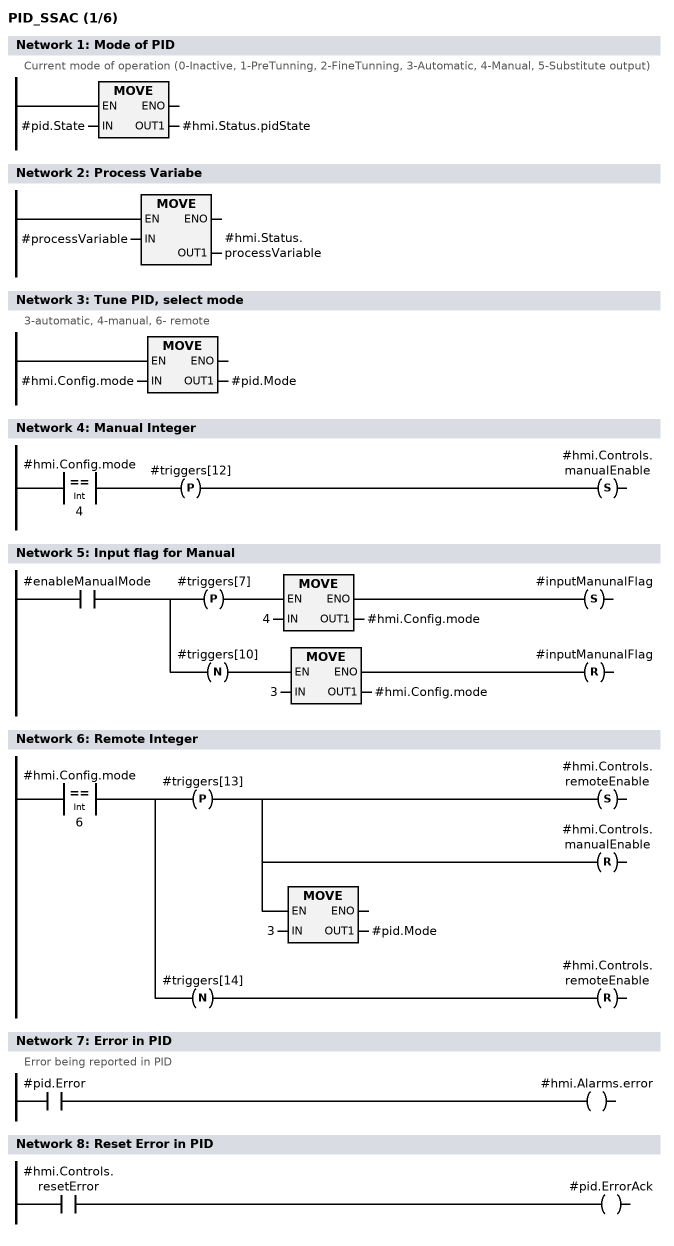
   RUNG wire#powerrail
      Move(in := #pid.State, out1 => #hmi.Status.pidState)
   END_RUNG
   // the same network as SCL:
   #hmi.Status.pidState := #pid.State;
END_REGION

REGION Network 2: Process Variabe
   RUNG wire#powerrail
      Move(in := #processVariable, out1 => #hmi.Status.processVariable)
   END_RUNG
   // the same network as SCL:
   #hmi.Status.processVariable := #processVariable;
END_REGION

REGION Network 3: Tune PID, select mode
   // 3-automatic, 4-manual, 6- remote
   RUNG wire#powerrail
      Move(in := #hmi.Config.mode, out1 => #pid.Mode)
   END_RUNG
   // the same network as SCL:
   #pid.Mode := #hmi.Config.mode;
END_REGION

REGION Network 4: Manual Integer
   RUNG wire#powerrail
      { S7_Templates := "SrcType := Int" } EQ_Contact(in1 := #hmi.Config.mode, in2 := 4)
      P_Trig( #triggers[12] )
      S_Coil( #hmi.Controls.manualEnable )
   END_RUNG
   // the same network as SCL:
   #_w1 := #hmi.Config.mode = 4;
   #_w2 := #_w1 AND NOT #triggers[12];   // rising edge
   #triggers[12] := #_w1;
   IF #_w2 THEN #hmi.Controls.manualEnable := TRUE; END_IF;
END_REGION

REGION Network 5: Input flag for Manual
   RUNG wire#powerrail
      Contact( #enableManualMode )
      wire#w1
      P_Trig( #triggers[7] )
      Move(in := 4, out1 => #hmi.Config.mode)
      S_Coil( #inputManunalFlag )
   END_RUNG
   RUNG wire#w1
      N_Trig( #triggers[10] )
      Move(in := 3, out1 => #hmi.Config.mode)
      R_Coil( #inputManunalFlag )
   END_RUNG
   // the same network as SCL:
   #_w1 := #enableManualMode AND NOT #triggers[7];   // rising edge
   #triggers[7] := #enableManualMode;
   IF #_w1 THEN
       #hmi.Config.mode := 4;
       #inputManunalFlag := TRUE;
   END_IF;
   #_w2 := NOT #enableManualMode AND #triggers[10];   // falling edge
   #triggers[10] := #enableManualMode;
   IF #_w2 THEN
       #hmi.Config.mode := 3;
       #inputManunalFlag := FALSE;
   END_IF;
END_REGION

REGION Network 6: Remote Integer
   RUNG wire#powerrail
      { S7_Templates := "SrcType := Int" } EQ_Contact(in1 := #hmi.Config.mode, in2 := 6)
      wire#w1
      P_Trig( #triggers[13] )
      wire#w2
      S_Coil( #hmi.Controls.remoteEnable )
   END_RUNG
   RUNG wire#w2
      R_Coil( #hmi.Controls.manualEnable )
   END_RUNG
   RUNG wire#w2
      Move(in := 3, out1 => #pid.Mode)
   END_RUNG
   RUNG wire#w1
      N_Trig( #triggers[14] )
      R_Coil( #hmi.Controls.remoteEnable )
   END_RUNG
   // the same network as SCL:
   #_w1 := #hmi.Config.mode = 6;
   #_w2 := #_w1 AND NOT #triggers[13];   // rising edge
   #triggers[13] := #_w1;
   IF #_w2 THEN
       #hmi.Controls.remoteEnable := TRUE;
       #hmi.Controls.manualEnable := FALSE;
       #pid.Mode := 3;
   END_IF;
   #_w3 := NOT #_w1 AND #triggers[14];   // falling edge
   #triggers[14] := #_w1;
   IF #_w3 THEN #hmi.Controls.remoteEnable := FALSE; END_IF;
END_REGION

REGION Network 7: Error in PID
   // Error being reported in PID
   RUNG wire#powerrail
      Contact( #pid.Error )
      Coil( #hmi.Alarms.error )
   END_RUNG
   // the same network as SCL:
   #hmi.Alarms.error := #pid.Error;
END_REGION

REGION Network 8: Reset Error in PID
   RUNG wire#powerrail
      Contact( #hmi.Controls.resetError )
      Coil( #pid.ErrorAck )
   END_RUNG
   // the same network as SCL:
   #pid.ErrorAck := #hmi.Controls.resetError;
END_REGION

REGION Network 9: Reset the controller if a change of Mode has been requested
   // mode 2 3 4 available thru here
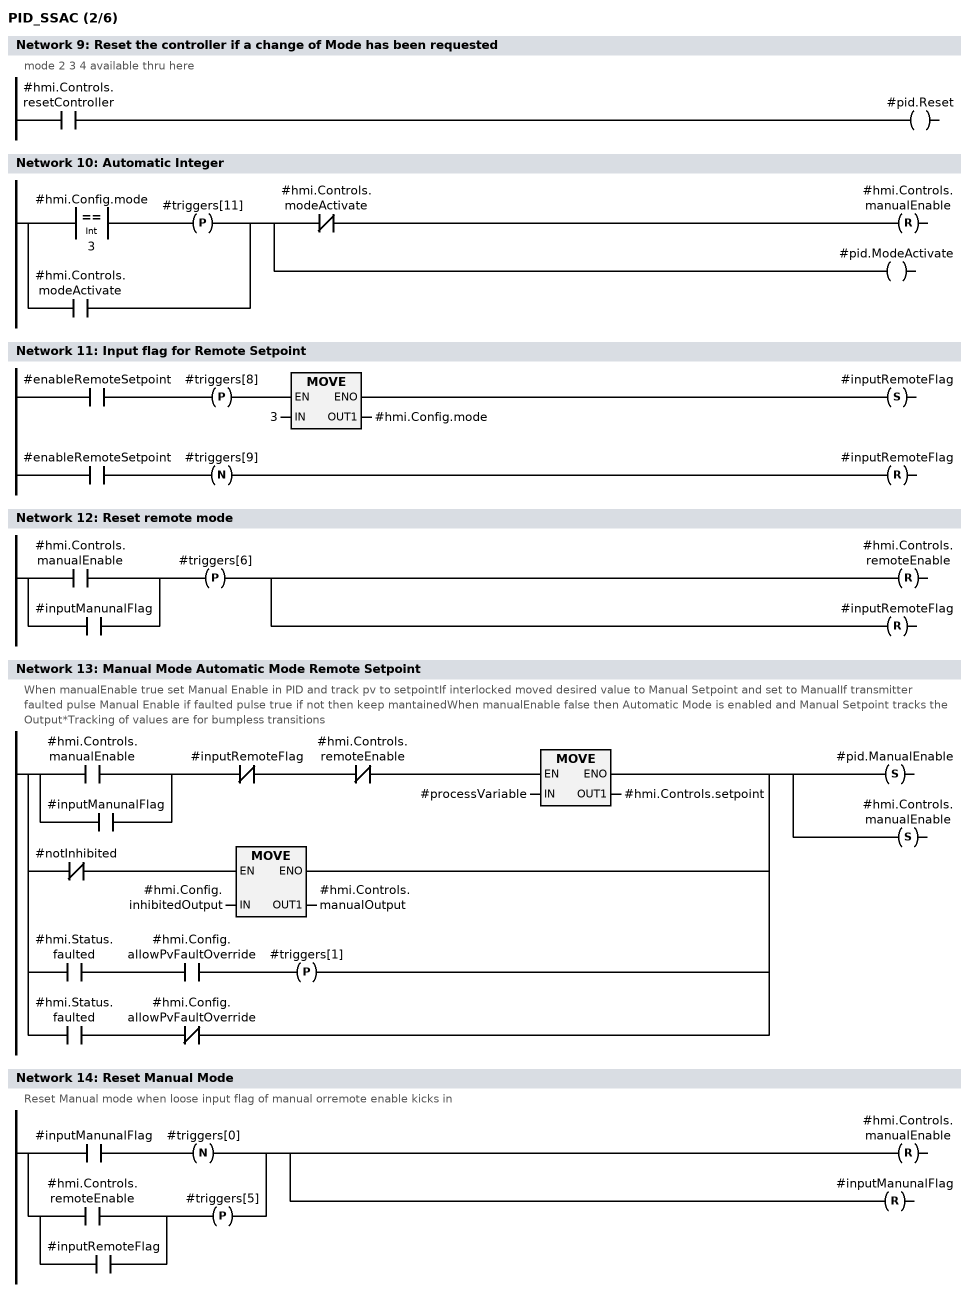
   RUNG wire#powerrail
      Contact( #hmi.Controls.resetController )
      Coil( #pid.Reset )
   END_RUNG
   // the same network as SCL:
   #pid.Reset := #hmi.Controls.resetController;
END_REGION

REGION Network 10: Automatic Integer
   RUNG wire#powerrail
      { S7_Templates := "SrcType := Int" } EQ_Contact(in1 := #hmi.Config.mode, in2 := 3)
      P_Trig( #triggers[11] )
      wire#w1
      I_Contact( #hmi.Controls.modeActivate )
      R_Coil( #hmi.Controls.manualEnable )
   END_RUNG
   RUNG wire#powerrail
      Contact( #hmi.Controls.modeActivate )
   END_RUNG wire#w1
   RUNG wire#w1
      Coil( #pid.ModeActivate )
   END_RUNG
   // the same network as SCL:
   #_w1 := #hmi.Config.mode = 3;
   #_w2 := #_w1 AND NOT #triggers[11];   // rising edge
   #triggers[11] := #_w1;
   #_w3 := #_w2 OR #hmi.Controls.modeActivate;
   IF #_w3 AND NOT #hmi.Controls.modeActivate THEN #hmi.Controls.manualEnable := FALSE; END_IF;
   #pid.ModeActivate := #_w3;
END_REGION

REGION Network 11: Input flag for Remote Setpoint
   RUNG wire#powerrail
      Contact( #enableRemoteSetpoint )
      P_Trig( #triggers[8] )
      Move(in := 3, out1 => #hmi.Config.mode)
      S_Coil( #inputRemoteFlag )
   END_RUNG
   RUNG wire#powerrail
      Contact( #enableRemoteSetpoint )
      N_Trig( #triggers[9] )
      R_Coil( #inputRemoteFlag )
   END_RUNG
   // the same network as SCL:
   #_w1 := #enableRemoteSetpoint AND NOT #triggers[8];   // rising edge
   #triggers[8] := #enableRemoteSetpoint;
   IF #_w1 THEN
       #hmi.Config.mode := 3;
       #inputRemoteFlag := TRUE;
   END_IF;
   #_w2 := NOT #enableRemoteSetpoint AND #triggers[9];   // falling edge
   #triggers[9] := #enableRemoteSetpoint;
   IF #_w2 THEN #inputRemoteFlag := FALSE; END_IF;
END_REGION

REGION Network 12: Reset remote mode
   RUNG wire#powerrail
      Contact( #hmi.Controls.manualEnable )
      wire#w1
      P_Trig( #triggers[6] )
      wire#w2
      R_Coil( #hmi.Controls.remoteEnable )
   END_RUNG
   RUNG wire#powerrail
      Contact( #inputManunalFlag )
   END_RUNG wire#w1
   RUNG wire#w2
      R_Coil( #inputRemoteFlag )
   END_RUNG
   // the same network as SCL:
   #_w1 := #hmi.Controls.manualEnable OR #inputManunalFlag;
   #_w2 := #_w1 AND NOT #triggers[6];   // rising edge
   #triggers[6] := #_w1;
   IF #_w2 THEN
       #hmi.Controls.remoteEnable := FALSE;
       #inputRemoteFlag := FALSE;
   END_IF;
END_REGION

REGION Network 13: Manual Mode Automatic Mode Remote Setpoint
   // When manualEnable true set Manual Enable in PID and track pv to setpointIf interlocked moved desired value to Manual Setpoint and set to ManualIf transmitter faulted pulse Manual Enable if faulted pulse true if not then keep mantainedWhen manualEnable false then Automatic Mode is enabled and Manual Setpoint tracks the Output*Tracking of values are for bumpless transitions
   RUNG wire#powerrail
      Contact( #hmi.Controls.manualEnable )
      wire#w1
      I_Contact( #inputRemoteFlag )
      I_Contact( #hmi.Controls.remoteEnable )
      Move(in := #processVariable, out1 => #hmi.Controls.setpoint)
      wire#w2
      S_Coil( #pid.ManualEnable )
   END_RUNG
   RUNG wire#powerrail
      Contact( #inputManunalFlag )
   END_RUNG wire#w1
   RUNG wire#powerrail
      I_Contact( #notInhibited )
      Move(in := #hmi.Config.inhibitedOutput, out1 => #hmi.Controls.manualOutput)
   END_RUNG wire#w2
   RUNG wire#powerrail
      Contact( #hmi.Status.faulted )
      Contact( #hmi.Config.allowPvFaultOverride )
      P_Trig( #triggers[1] )
   END_RUNG wire#w2
   RUNG wire#powerrail
      Contact( #hmi.Status.faulted )
      I_Contact( #hmi.Config.allowPvFaultOverride )
   END_RUNG wire#w2
   RUNG wire#w2
      S_Coil( #hmi.Controls.manualEnable )
   END_RUNG
   // the same network as SCL:
   #_w1 := (#hmi.Controls.manualEnable OR #inputManunalFlag) AND NOT #inputRemoteFlag AND NOT #hmi.Controls.remoteEnable;
   IF #_w1 THEN #hmi.Controls.setpoint := #processVariable; END_IF;
   IF NOT #notInhibited THEN #hmi.Controls.manualOutput := #hmi.Config.inhibitedOutput; END_IF;
   #_w2 := #hmi.Status.faulted AND #hmi.Config.allowPvFaultOverride;
   #_w3 := #_w2 AND NOT #triggers[1];   // rising edge
   #triggers[1] := #_w2;
   IF #_w1 OR NOT #notInhibited OR #_w3 OR (#hmi.Status.faulted AND NOT #hmi.Config.allowPvFaultOverride) THEN
       #pid.ManualEnable := TRUE;
       #hmi.Controls.manualEnable := TRUE;
   END_IF;
END_REGION

REGION Network 14: Reset Manual Mode
   // Reset Manual mode when loose input flag of manual orremote enable kicks in
   RUNG wire#powerrail
      Contact( #inputManunalFlag )
      N_Trig( #triggers[0] )
      wire#w1
      R_Coil( #hmi.Controls.manualEnable )
   END_RUNG
   RUNG wire#powerrail
      Contact( #hmi.Controls.remoteEnable )
      wire#w2
      P_Trig( #triggers[5] )
   END_RUNG wire#w1
   RUNG wire#powerrail
      Contact( #inputRemoteFlag )
   END_RUNG wire#w2
   RUNG wire#w1
      R_Coil( #inputManunalFlag )
   END_RUNG
   // the same network as SCL:
   #_w1 := NOT #inputManunalFlag AND #triggers[0];   // falling edge
   #triggers[0] := #inputManunalFlag;
   #_w2 := #hmi.Controls.remoteEnable OR #inputRemoteFlag;
   #_w3 := #_w2 AND NOT #triggers[5];   // rising edge
   #triggers[5] := #_w2;
   IF #_w1 OR #_w3 THEN
       #hmi.Controls.manualEnable := FALSE;
       #inputManunalFlag := FALSE;
   END_IF;
END_REGION

REGION Network 15: Automatic Mode
   // IF not in manual and not in remote then in Automatic mode, reset Manual Mode of  PID
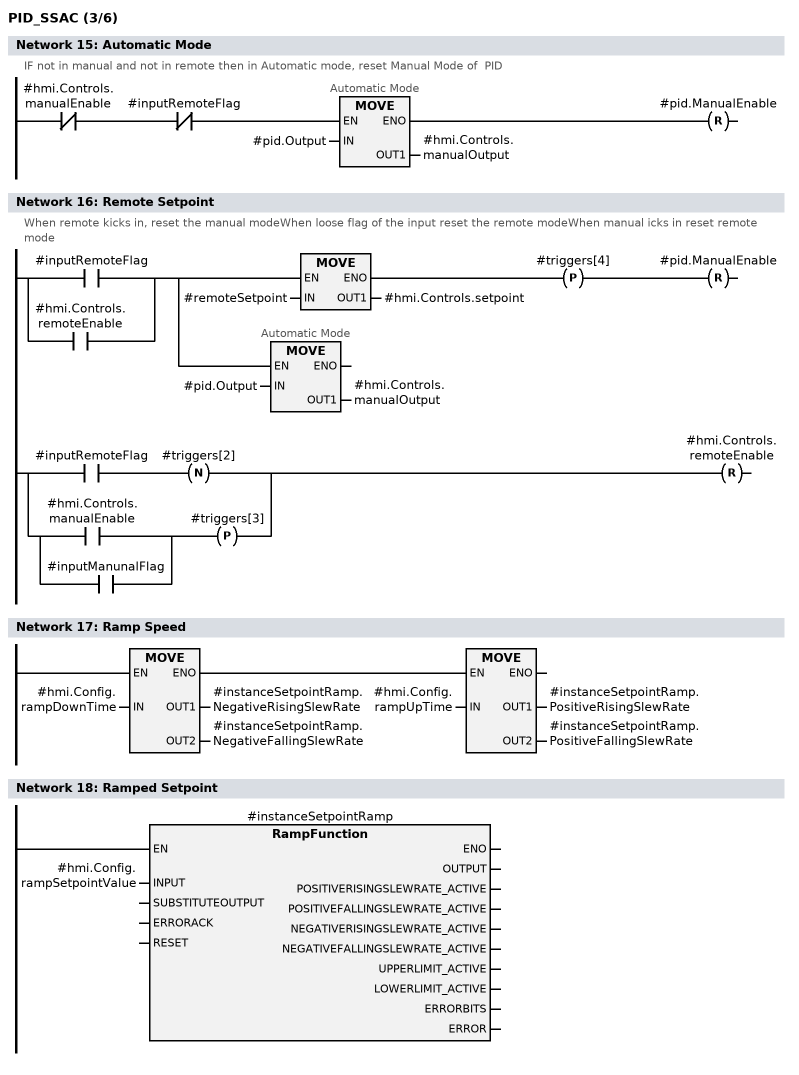
   RUNG wire#powerrail
      I_Contact( #hmi.Controls.manualEnable )
      I_Contact( #inputRemoteFlag )
      Move(in := #pid.Output, out1 => #hmi.Controls.manualOutput)   // Automatic Mode
      R_Coil( #pid.ManualEnable )
   END_RUNG
   // the same network as SCL:
   IF NOT #hmi.Controls.manualEnable AND NOT #inputRemoteFlag THEN
       #hmi.Controls.manualOutput := #pid.Output;   // Automatic Mode
       #pid.ManualEnable := FALSE;
   END_IF;
END_REGION

REGION Network 16: Remote Setpoint
   // When remote kicks in, reset the manual modeWhen loose flag of the input reset the remote modeWhen manual icks in reset remote mode
   RUNG wire#powerrail
      Contact( #inputRemoteFlag )
      wire#w1
      Move(in := #remoteSetpoint, out1 => #hmi.Controls.setpoint)
      P_Trig( #triggers[4] )
      R_Coil( #pid.ManualEnable )
   END_RUNG
   RUNG wire#powerrail
      Contact( #hmi.Controls.remoteEnable )
   END_RUNG wire#w1
   RUNG wire#w1
      Move(in := #pid.Output, out1 => #hmi.Controls.manualOutput)   // Automatic Mode
   END_RUNG
   RUNG wire#powerrail
      Contact( #inputRemoteFlag )
      N_Trig( #triggers[2] )
      wire#w2
      R_Coil( #hmi.Controls.remoteEnable )
   END_RUNG
   RUNG wire#powerrail
      Contact( #hmi.Controls.manualEnable )
      wire#w3
      P_Trig( #triggers[3] )
   END_RUNG wire#w2
   RUNG wire#powerrail
      Contact( #inputManunalFlag )
   END_RUNG wire#w3
   // the same network as SCL:
   #_w1 := #inputRemoteFlag OR #hmi.Controls.remoteEnable;
   IF #_w1 THEN #hmi.Controls.setpoint := #remoteSetpoint; END_IF;
   #_w2 := #_w1 AND NOT #triggers[4];   // rising edge
   #triggers[4] := #_w1;
   IF #_w2 THEN #pid.ManualEnable := FALSE; END_IF;
   IF #_w1 THEN
       #hmi.Controls.manualOutput := #pid.Output;   // Automatic Mode
   END_IF;
   #_w3 := NOT #inputRemoteFlag AND #triggers[2];   // falling edge
   #triggers[2] := #inputRemoteFlag;
   #_w4 := #hmi.Controls.manualEnable OR #inputManunalFlag;
   #_w5 := #_w4 AND NOT #triggers[3];   // rising edge
   #triggers[3] := #_w4;
   IF #_w3 OR #_w5 THEN #hmi.Controls.remoteEnable := FALSE; END_IF;
END_REGION

REGION Network 17: Ramp Speed
   RUNG wire#powerrail
      Move(in := #hmi.Config.rampDownTime, out1 => #instanceSetpointRamp.NegativeRisingSlewRate, out2 => #instanceSetpointRamp.NegativeFallingSlewRate)
      Move(in := #hmi.Config.rampUpTime, out1 => #instanceSetpointRamp.PositiveRisingSlewRate, out2 => #instanceSetpointRamp.PositiveFallingSlewRate)
   END_RUNG
   // the same network as SCL:
   #instanceSetpointRamp.NegativeRisingSlewRate := #hmi.Config.rampDownTime;
   #instanceSetpointRamp.NegativeFallingSlewRate := #hmi.Config.rampDownTime;
   #instanceSetpointRamp.PositiveRisingSlewRate := #hmi.Config.rampUpTime;
   #instanceSetpointRamp.PositiveFallingSlewRate := #hmi.Config.rampUpTime;
END_REGION

REGION Network 18: Ramped Setpoint
   #instanceSetpointRamp(Input := #hmi.Config.rampSetpointValue);   // RampFunction
END_REGION

REGION Network 19: Setpoint Control
   // If ramp enabled then move ramped setpointif ramp disabled then move hmi setpoint
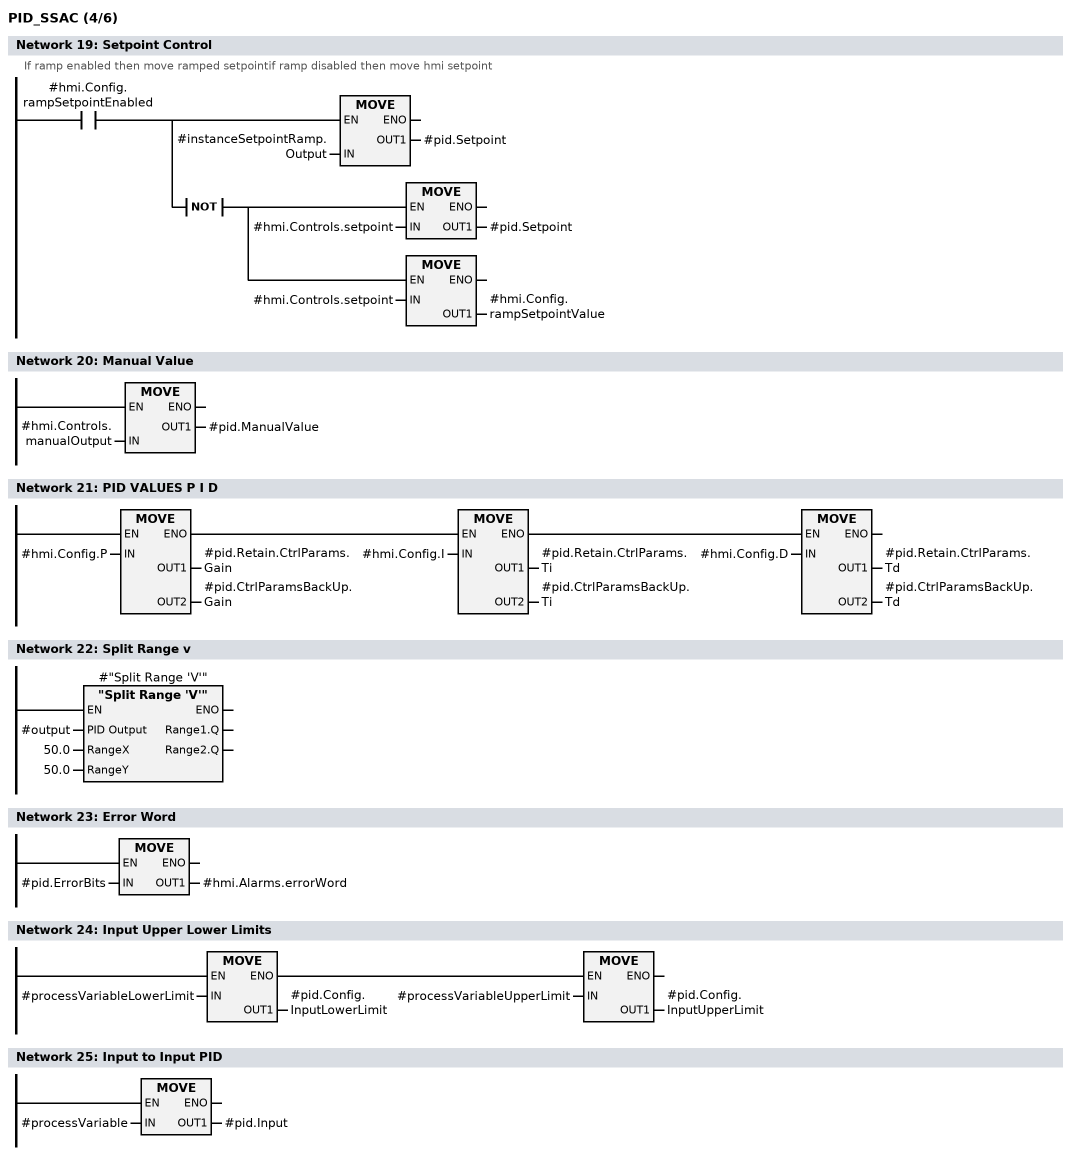
   RUNG wire#powerrail
      Contact( #hmi.Config.rampSetpointEnabled )
      wire#w1
      Move(in := #instanceSetpointRamp.Output, out1 => #pid.Setpoint)
   END_RUNG
   RUNG wire#w1
      Not()
      wire#w2
      Move(in := #hmi.Controls.setpoint, out1 => #pid.Setpoint)
   END_RUNG
   RUNG wire#w2
      Move(in := #hmi.Controls.setpoint, out1 => #hmi.Config.rampSetpointValue)
   END_RUNG
   // the same network as SCL:
   IF #hmi.Config.rampSetpointEnabled THEN #pid.Setpoint := #instanceSetpointRamp.Output; END_IF;
   IF NOT #hmi.Config.rampSetpointEnabled THEN
       #pid.Setpoint := #hmi.Controls.setpoint;
       #hmi.Config.rampSetpointValue := #hmi.Controls.setpoint;
   END_IF;
END_REGION

REGION Network 20: Manual Value
   RUNG wire#powerrail
      Move(in := #hmi.Controls.manualOutput, out1 => #pid.ManualValue)
   END_RUNG
   // the same network as SCL:
   #pid.ManualValue := #hmi.Controls.manualOutput;
END_REGION

REGION Network 21: PID VALUES P I D
   RUNG wire#powerrail
      Move(in := #hmi.Config.P, out1 => #pid.Retain.CtrlParams.Gain, out2 => #pid.CtrlParamsBackUp.Gain)
      Move(in := #hmi.Config.I, out1 => #pid.Retain.CtrlParams.Ti, out2 => #pid.CtrlParamsBackUp.Ti)
      Move(in := #hmi.Config.D, out1 => #pid.Retain.CtrlParams.Td, out2 => #pid.CtrlParamsBackUp.Td)
   END_RUNG
   // the same network as SCL:
   #pid.Retain.CtrlParams.Gain := #hmi.Config.P;
   #pid.CtrlParamsBackUp.Gain := #hmi.Config.P;
   #pid.Retain.CtrlParams.Ti := #hmi.Config.I;
   #pid.CtrlParamsBackUp.Ti := #hmi.Config.I;
   #pid.Retain.CtrlParams.Td := #hmi.Config.D;
   #pid.CtrlParamsBackUp.Td := #hmi.Config.D;
END_REGION

REGION Network 22: Split Range v
   RUNG wire#powerrail
      #"Split Range 'V'"("PID Output" := #output, RangeX := 50.0, RangeY := 50.0, "Range1.Q" =>, "Range2.Q" =>)
   END_RUNG
   // the same network as SCL:
   #"Split Range 'V'"("PID Output" := #output, RangeX := 50.0, RangeY := 50.0);   // "Split Range 'V'"
END_REGION

REGION Network 23: Error Word
   RUNG wire#powerrail
      Move(in := #pid.ErrorBits, out1 => #hmi.Alarms.errorWord)
   END_RUNG
   // the same network as SCL:
   #hmi.Alarms.errorWord := #pid.ErrorBits;
END_REGION

REGION Network 24: Input Upper Lower Limits
   RUNG wire#powerrail
      Move(in := #processVariableLowerLimit, out1 => #pid.Config.InputLowerLimit)
      Move(in := #processVariableUpperLimit, out1 => #pid.Config.InputUpperLimit)
   END_RUNG
   // the same network as SCL:
   #pid.Config.InputLowerLimit := #processVariableLowerLimit;
   #pid.Config.InputUpperLimit := #processVariableUpperLimit;
END_REGION

REGION Network 25: Input to Input PID
   RUNG wire#powerrail
      Move(in := #processVariable, out1 => #pid.Input)
   END_RUNG
   // the same network as SCL:
   #pid.Input := #processVariable;
END_REGION

REGION Network 26: Outputs
   // Outputs of PID block
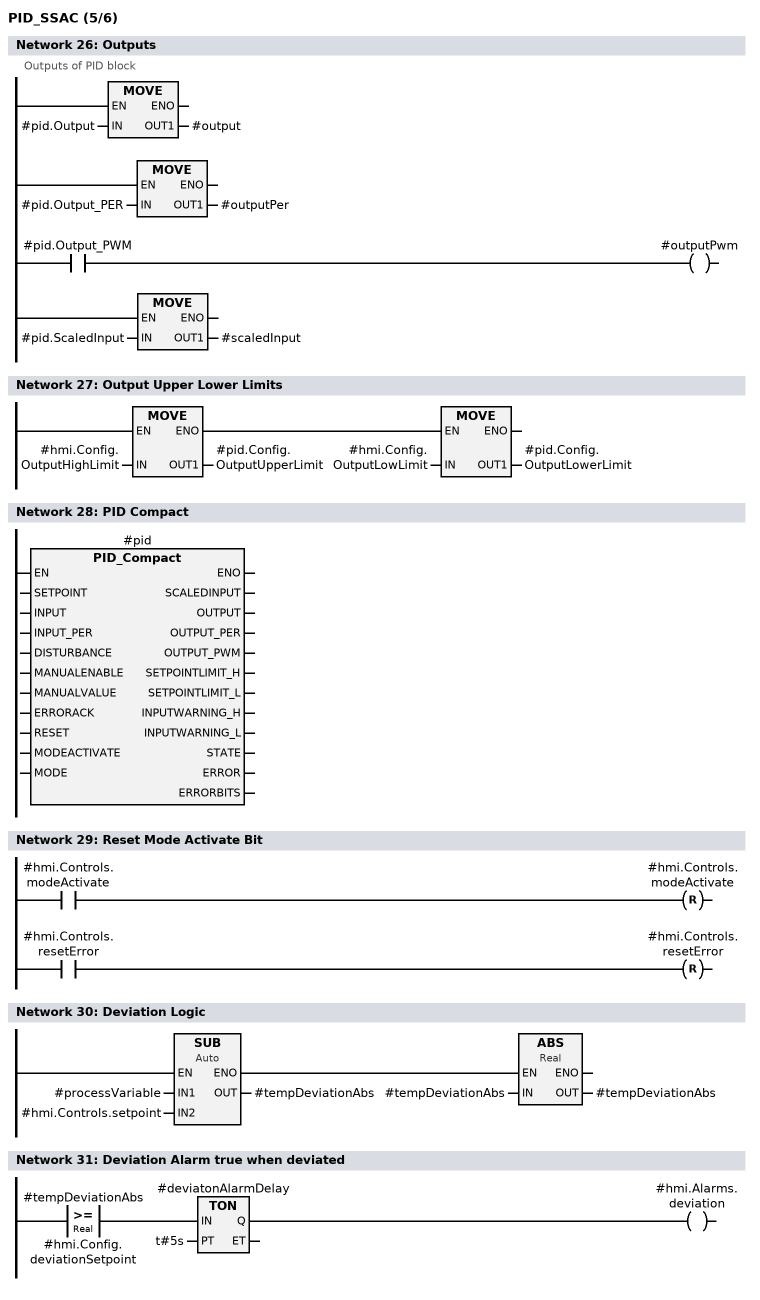
   RUNG wire#powerrail
      Move(in := #pid.Output, out1 => #output)
   END_RUNG
   RUNG wire#powerrail
      Move(in := #pid.Output_PER, out1 => #outputPer)
   END_RUNG
   RUNG wire#powerrail
      Contact( #pid.Output_PWM )
      Coil( #outputPwm )
   END_RUNG
   RUNG wire#powerrail
      Move(in := #pid.ScaledInput, out1 => #scaledInput)
   END_RUNG
   // the same network as SCL:
   #output := #pid.Output;
   #outputPer := #pid.Output_PER;
   #outputPwm := #pid.Output_PWM;
   #scaledInput := #pid.ScaledInput;
END_REGION

REGION Network 27: Output Upper Lower Limits
   RUNG wire#powerrail
      Move(in := #hmi.Config.OutputHighLimit, out1 => #pid.Config.OutputUpperLimit)
      Move(in := #hmi.Config.OutputLowLimit, out1 => #pid.Config.OutputLowerLimit)
   END_RUNG
   // the same network as SCL:
   #pid.Config.OutputUpperLimit := #hmi.Config.OutputHighLimit;
   #pid.Config.OutputLowerLimit := #hmi.Config.OutputLowLimit;
END_REGION

REGION Network 28: PID Compact
   #pid();   // PID_Compact
END_REGION

REGION Network 29: Reset Mode Activate Bit
   RUNG wire#powerrail
      Contact( #hmi.Controls.modeActivate )
      R_Coil( #hmi.Controls.modeActivate )
   END_RUNG
   RUNG wire#powerrail
      Contact( #hmi.Controls.resetError )
      R_Coil( #hmi.Controls.resetError )
   END_RUNG
   // the same network as SCL:
   IF #hmi.Controls.modeActivate THEN #hmi.Controls.modeActivate := FALSE; END_IF;
   IF #hmi.Controls.resetError THEN #hmi.Controls.resetError := FALSE; END_IF;
END_REGION

REGION Network 30: Deviation Logic
   RUNG wire#powerrail
      Sub(in1 := #processVariable, in2 := #hmi.Controls.setpoint, out => #tempDeviationAbs)
      { S7_Templates := "SrcType := Real" } Abs(in := #tempDeviationAbs, out => #tempDeviationAbs)
   END_RUNG
   // the same network as SCL:
   #tempDeviationAbs := #processVariable - #hmi.Controls.setpoint;
   #tempDeviationAbs := ABS(#tempDeviationAbs);
END_REGION

REGION Network 31: Deviation Alarm true when deviated
   #deviatonAlarmDelay(IN := #tempDeviationAbs >= #hmi.Config.deviationSetpoint, PT := t#5s);   // TON
   #hmi.Alarms.deviation := #deviatonAlarmDelay.Q;
END_REGION

REGION Network 32: PID inhibited (interlocked, off)
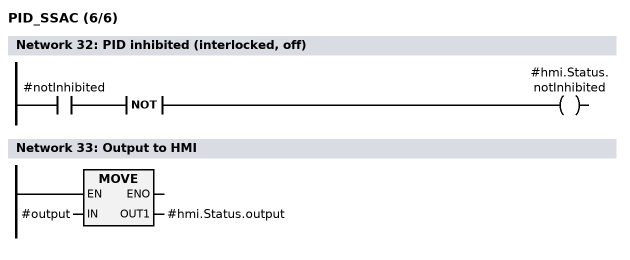
   RUNG wire#powerrail
      Contact( #notInhibited )
      Not()
      Coil( #hmi.Status.notInhibited )
   END_RUNG
   // the same network as SCL:
   #hmi.Status.notInhibited := NOT #notInhibited;
END_REGION

REGION Network 33: Output to HMI
   RUNG wire#powerrail
      Move(in := #output, out1 => #hmi.Status.output)
   END_RUNG
   // the same network as SCL:
   #hmi.Status.output := #output;
END_REGION
END_FUNCTION_BLOCK

FUNCTION_BLOCK "Totalizer_Siemens"   // FB3, SCL
{ S7_Optimized_Access := 'TRUE' }
VERSION : 0.1
   VAR_INPUT
      value : Real;
      intervall : Time;
      cycle : Time;
      reset : Bool;
   END_VAR
   VAR_OUTPUT
      total : Real;
   END_VAR
   VAR
      statAccum : Real;
   END_VAR
   VAR_TEMP
      tempIntervall : Real;
      tempCycle : Real;
      tempIntervallDInt : DInt;
      tempCycleDInt : DInt;
   END_VAR
BEGIN
   //Ist der Signalzustand der Variable "Reset" gleich True, so werden die Variablen
   //"Accum" und "Total" auf Null zurückgesetzt und es erfolgt keine Berechnung.
   //Beim Signalzustand False erfolgt zunächst eine Datentypumwandlung nach Real der beiden
   //Eingangsvariablen "Intervall" und "Cycle". Zuerst mit der Konvertierung von Time nach
   //DInt und anschließend von DInt nach Real.
   //Innerhalb eines Zyklus wird der Eingangswert der Variablen "Value" mit dem Wert der temporären Variablen
   //"Cycle_real" multipliziert und mit dem Wert der temporären Variablen "Intervall_real" dividiert.
   //Das Ergebnis wird anschließend in den Zwischenspeicher "Accum" abgelegt. Somit wird innerhalb eines jeden
   //Zykluses das Zwischenergebnis im "Accum" um diesen Wert inkrementiert, welches auch in jedem Zyklus zur
   //Ausgangsvariable "Total" transferiert wird.
   //***************************************************************************
   //If the signal status of the variable "Reset" is true, the variables "Accum" and "Total"
   //are set to zero and there is no calculation.
   //If the signal status is false, there is first a data type change to real of the two
   //input variables "Intervall" and "Cycle. After conversion from Time to DInit and from DInt to Real.
   //In a #Cycle the input #Value of the variable "Value" is multiplied by the #Value of the temporary variable
   //"Cycle_real" and then divided by the #Value of the temporary variable "Intervall_real". The result is then
   //stored in the buffer "Accum". This in one particular #Cycle the result in the "Accum" buffer is
   //incremented this #Value, which is also transferred to the output variable "Total" in that #Cycle too.

   IF #reset = true THEN
       #statAccum := 0.000000e000; //Die Variablen werden zurückgesetzt.
       #total := 0.000000e000; //The variables will be set to zero.
   ELSE
       #tempIntervallDInt := TIME_TO_DINT(#intervall);
       #tempIntervall := DINT_TO_REAL(#tempIntervallDInt);
       #tempCycleDInt := TIME_TO_DINT(#cycle);
       #tempCycle := DINT_TO_REAL(#tempCycleDInt);
       #statAccum := ((#value * #tempCycle) / #tempIntervall) + #statAccum;
       #total := #statAccum; //Kopiere Ergebnis nach #Total / Copy result to #Total.
   END_IF;
END_FUNCTION_BLOCK

FUNCTION_BLOCK "PID_TIA"   // FB814, LAD
{ S7_Optimized_Access := 'TRUE' }
VERSION : 0.1
   VAR_INPUT
      processVariable : Real;
      processVariableLowerLimit : Real;
      processVariableUpperLimit : Real;
      notInhibited : Bool := TRUE;
      remoteSetpoint : Real;
      enableManualMode : Bool;
      enableRemoteSetpoint : Bool;
   END_VAR
   VAR_OUTPUT
      scaledInput : Real;
      output : Real;   // Manipulated Value REAL
      outputPer : Int;   // Manipulated Value INT
      outputPwm : Bool;   // Output PWM
   END_VAR
   VAR_IN_OUT
      pid : PID_Compact;
   END_VAR
   VAR
      hmi : Struct
         Controls : Struct
            setpoint : Real;   // Setpoint sent to PID
            manualEnable : Bool;   // Enables Manual mode
            manualOutput : Real;   // Manual Output sent to PID 0 to 100 %
            remoteEnable : Bool;
            resetController : Bool;   // Resets Controller sent to PID
            resetError : Bool;   // ErrorAck to PID
            modeActivate : Bool;   // Execute the change of mode
         END_STRUCT;
         Config : Struct
            P : Real := 0.1;   // Proportional Control sent to PID
            I : Real := 10.0;   // Integral Control sent to PID
            D : Real := 0.0;   // Derivative Control sent to PID
            OutputHighLimit : Real := 100.0;   // Output Upper Limit sent to PID
            OutputLowLimit : Real := 0.0;   // Output Lower Limit sent to PID
            rampDownTime : Real := 1.0;
            rampUpTime : Real := 1.0;
            allowPvFaultOverride : Bool;   // Allows operator to override PV fault
            rampSetpointEnabled : Bool;   // Enables the ramping of a setpoint inside the PID
            rampSetpointValue : Real;   // Value to be reached in the ramp
            inhibitedOutput : Real := 0.0;   // Inhibited Value set by the Operator 0 to 100
            mode : Int := 4;   // Mode selected by operator 1=pretune,2=finetuning,3=automatic,4-manual, 5-Substitute output, 6-Remote
            enablePVtracking : Bool;
         END_STRUCT;
         Status : Struct
            faulted : Bool;   // Transmitter Faulted
            notInhibited : Bool;   // PID inhibited (interlocked, off)
            pidState : Int;   // Current mode of operation (0-Inactive, 1-SUT, 2-TIR, 3-Automatic, 4-Manual, 5-Substitute output)
            Output : Real;   // Output of the PID
         END_STRUCT;
         Alarms : Struct
            errorWord : DWord;   // Error Word of PID
            error : Bool;   // Error in PID
         END_STRUCT;
      END_STRUCT;
      triggers : Array[0..20] of Bool;
      inputManunalFlag : Bool;
      inputRemoteFlag : Bool;
      "Dont Overwrite SP" : Bool;
      trig : Bool;
      trig2 : Bool;
      trig3 : Bool;
      "Let ramp" : Bool;
      IEC_Timer_0_Instance : TON_TIME;
      Ramp_Instance : "Ramp";
   END_VAR
   VAR_TEMP
      tempIgnore : Bool;
   END_VAR
   VAR_TEMP   // added for the SCL form of the ladder/FBD networks
      _w1 : Bool;
      _w2 : Bool;
      _w3 : Bool;
      _w4 : Bool;
      _w5 : Bool;
   END_VAR
BEGIN

REGION Network 1: PID inhibited (interlocked, off)
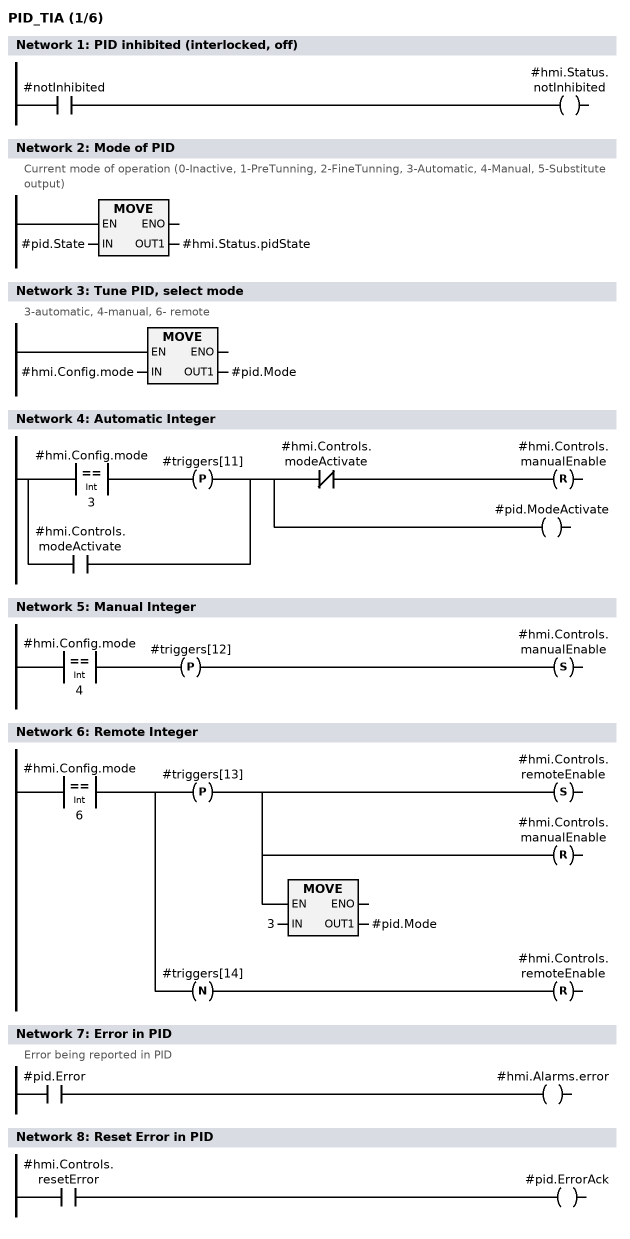
   RUNG wire#powerrail
      Contact( #notInhibited )
      Coil( #hmi.Status.notInhibited )
   END_RUNG
   // the same network as SCL:
   #hmi.Status.notInhibited := #notInhibited;
END_REGION

REGION Network 2: Mode of PID
   // Current mode of operation (0-Inactive, 1-PreTunning, 2-FineTunning, 3-Automatic, 4-Manual, 5-Substitute output)
   RUNG wire#powerrail
      Move(in := #pid.State, out1 => #hmi.Status.pidState)
   END_RUNG
   // the same network as SCL:
   #hmi.Status.pidState := #pid.State;
END_REGION

REGION Network 3: Tune PID, select mode
   // 3-automatic, 4-manual, 6- remote
   RUNG wire#powerrail
      Move(in := #hmi.Config.mode, out1 => #pid.Mode)
   END_RUNG
   // the same network as SCL:
   #pid.Mode := #hmi.Config.mode;
END_REGION

REGION Network 4: Automatic Integer
   RUNG wire#powerrail
      { S7_Templates := "SrcType := Int" } EQ_Contact(in1 := #hmi.Config.mode, in2 := 3)
      P_Trig( #triggers[11] )
      wire#w1
      I_Contact( #hmi.Controls.modeActivate )
      R_Coil( #hmi.Controls.manualEnable )
   END_RUNG
   RUNG wire#powerrail
      Contact( #hmi.Controls.modeActivate )
   END_RUNG wire#w1
   RUNG wire#w1
      Coil( #pid.ModeActivate )
   END_RUNG
   // the same network as SCL:
   #_w1 := #hmi.Config.mode = 3;
   #_w2 := #_w1 AND NOT #triggers[11];   // rising edge
   #triggers[11] := #_w1;
   #_w3 := #_w2 OR #hmi.Controls.modeActivate;
   IF #_w3 AND NOT #hmi.Controls.modeActivate THEN #hmi.Controls.manualEnable := FALSE; END_IF;
   #pid.ModeActivate := #_w3;
END_REGION

REGION Network 5: Manual Integer
   RUNG wire#powerrail
      { S7_Templates := "SrcType := Int" } EQ_Contact(in1 := #hmi.Config.mode, in2 := 4)
      P_Trig( #triggers[12] )
      S_Coil( #hmi.Controls.manualEnable )
   END_RUNG
   // the same network as SCL:
   #_w1 := #hmi.Config.mode = 4;
   #_w2 := #_w1 AND NOT #triggers[12];   // rising edge
   #triggers[12] := #_w1;
   IF #_w2 THEN #hmi.Controls.manualEnable := TRUE; END_IF;
END_REGION

REGION Network 6: Remote Integer
   RUNG wire#powerrail
      { S7_Templates := "SrcType := Int" } EQ_Contact(in1 := #hmi.Config.mode, in2 := 6)
      wire#w1
      P_Trig( #triggers[13] )
      wire#w2
      S_Coil( #hmi.Controls.remoteEnable )
   END_RUNG
   RUNG wire#w2
      R_Coil( #hmi.Controls.manualEnable )
   END_RUNG
   RUNG wire#w2
      Move(in := 3, out1 => #pid.Mode)
   END_RUNG
   RUNG wire#w1
      N_Trig( #triggers[14] )
      R_Coil( #hmi.Controls.remoteEnable )
   END_RUNG
   // the same network as SCL:
   #_w1 := #hmi.Config.mode = 6;
   #_w2 := #_w1 AND NOT #triggers[13];   // rising edge
   #triggers[13] := #_w1;
   IF #_w2 THEN
       #hmi.Controls.remoteEnable := TRUE;
       #hmi.Controls.manualEnable := FALSE;
       #pid.Mode := 3;
   END_IF;
   #_w3 := NOT #_w1 AND #triggers[14];   // falling edge
   #triggers[14] := #_w1;
   IF #_w3 THEN #hmi.Controls.remoteEnable := FALSE; END_IF;
END_REGION

REGION Network 7: Error in PID
   // Error being reported in PID
   RUNG wire#powerrail
      Contact( #pid.Error )
      Coil( #hmi.Alarms.error )
   END_RUNG
   // the same network as SCL:
   #hmi.Alarms.error := #pid.Error;
END_REGION

REGION Network 8: Reset Error in PID
   RUNG wire#powerrail
      Contact( #hmi.Controls.resetError )
      Coil( #pid.ErrorAck )
   END_RUNG
   // the same network as SCL:
   #pid.ErrorAck := #hmi.Controls.resetError;
END_REGION

REGION Network 9: Reset the controller if a change of Mode has been requested
   // mode 2 3 4 available thru here
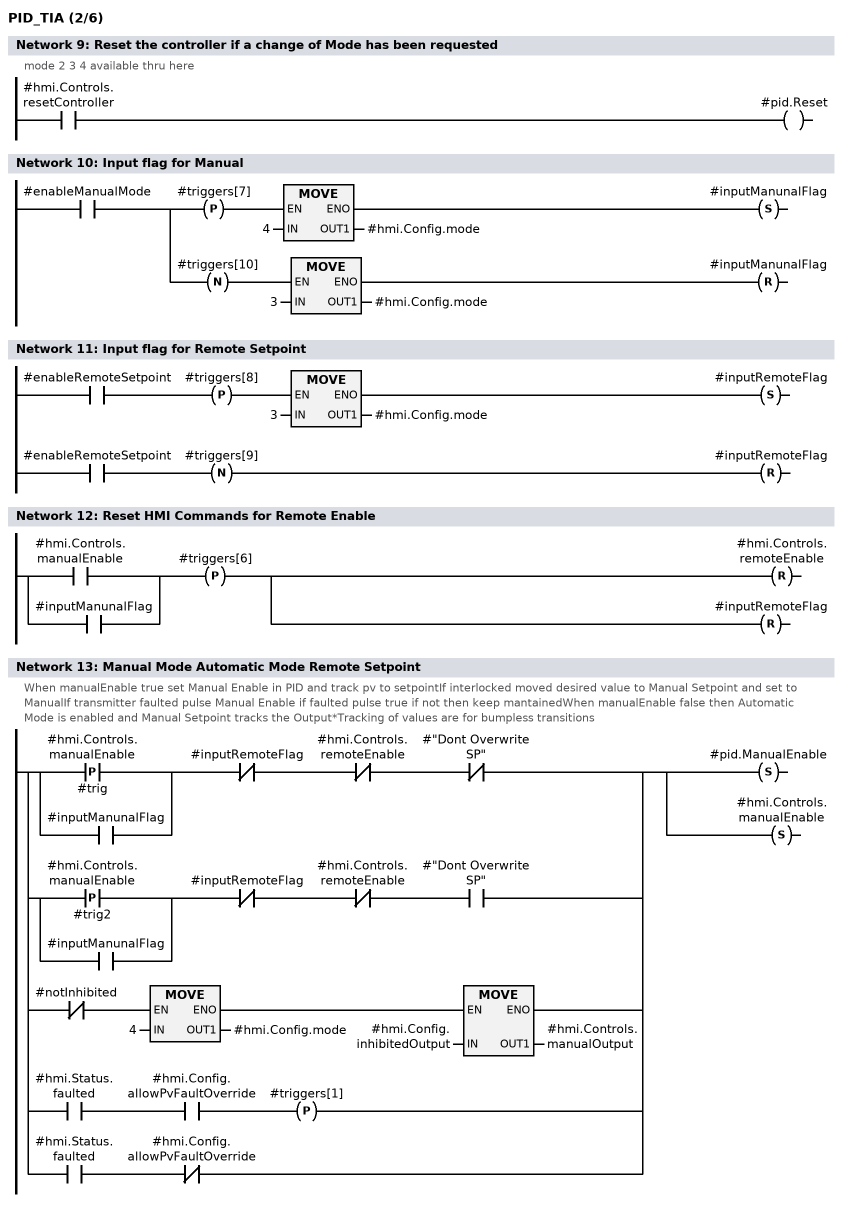
   RUNG wire#powerrail
      Contact( #hmi.Controls.resetController )
      Coil( #pid.Reset )
   END_RUNG
   // the same network as SCL:
   #pid.Reset := #hmi.Controls.resetController;
END_REGION

REGION Network 10: Input flag for Manual
   RUNG wire#powerrail
      Contact( #enableManualMode )
      wire#w1
      P_Trig( #triggers[7] )
      Move(in := 4, out1 => #hmi.Config.mode)
      S_Coil( #inputManunalFlag )
   END_RUNG
   RUNG wire#w1
      N_Trig( #triggers[10] )
      Move(in := 3, out1 => #hmi.Config.mode)
      R_Coil( #inputManunalFlag )
   END_RUNG
   // the same network as SCL:
   #_w1 := #enableManualMode AND NOT #triggers[7];   // rising edge
   #triggers[7] := #enableManualMode;
   IF #_w1 THEN
       #hmi.Config.mode := 4;
       #inputManunalFlag := TRUE;
   END_IF;
   #_w2 := NOT #enableManualMode AND #triggers[10];   // falling edge
   #triggers[10] := #enableManualMode;
   IF #_w2 THEN
       #hmi.Config.mode := 3;
       #inputManunalFlag := FALSE;
   END_IF;
END_REGION

REGION Network 11: Input flag for Remote Setpoint
   RUNG wire#powerrail
      Contact( #enableRemoteSetpoint )
      P_Trig( #triggers[8] )
      Move(in := 3, out1 => #hmi.Config.mode)
      S_Coil( #inputRemoteFlag )
   END_RUNG
   RUNG wire#powerrail
      Contact( #enableRemoteSetpoint )
      N_Trig( #triggers[9] )
      R_Coil( #inputRemoteFlag )
   END_RUNG
   // the same network as SCL:
   #_w1 := #enableRemoteSetpoint AND NOT #triggers[8];   // rising edge
   #triggers[8] := #enableRemoteSetpoint;
   IF #_w1 THEN
       #hmi.Config.mode := 3;
       #inputRemoteFlag := TRUE;
   END_IF;
   #_w2 := NOT #enableRemoteSetpoint AND #triggers[9];   // falling edge
   #triggers[9] := #enableRemoteSetpoint;
   IF #_w2 THEN #inputRemoteFlag := FALSE; END_IF;
END_REGION

REGION Network 12: Reset HMI Commands for Remote Enable
   RUNG wire#powerrail
      Contact( #hmi.Controls.manualEnable )
      wire#w1
      P_Trig( #triggers[6] )
      wire#w2
      R_Coil( #hmi.Controls.remoteEnable )
   END_RUNG
   RUNG wire#powerrail
      Contact( #inputManunalFlag )
   END_RUNG wire#w1
   RUNG wire#w2
      R_Coil( #inputRemoteFlag )
   END_RUNG
   // the same network as SCL:
   #_w1 := #hmi.Controls.manualEnable OR #inputManunalFlag;
   #_w2 := #_w1 AND NOT #triggers[6];   // rising edge
   #triggers[6] := #_w1;
   IF #_w2 THEN
       #hmi.Controls.remoteEnable := FALSE;
       #inputRemoteFlag := FALSE;
   END_IF;
END_REGION

REGION Network 13: Manual Mode Automatic Mode Remote Setpoint
   // When manualEnable true set Manual Enable in PID and track pv to setpointIf interlocked moved desired value to Manual Setpoint and set to ManualIf transmitter faulted pulse Manual Enable if faulted pulse true if not then keep mantainedWhen manualEnable false then Automatic Mode is enabled and Manual Setpoint tracks the Output*Tracking of values are for bumpless transitions
   RUNG wire#powerrail
      P_Contact(operand := #hmi.Controls.manualEnable, bit := #trig)
      wire#w1
      I_Contact( #inputRemoteFlag )
      I_Contact( #hmi.Controls.remoteEnable )
      I_Contact( #"Dont Overwrite SP" )
      wire#w2
      S_Coil( #pid.ManualEnable )
   END_RUNG
   RUNG wire#powerrail
      Contact( #inputManunalFlag )
   END_RUNG wire#w1
   RUNG wire#powerrail
      P_Contact(operand := #hmi.Controls.manualEnable, bit := #trig2)
      wire#w3
      I_Contact( #inputRemoteFlag )
      I_Contact( #hmi.Controls.remoteEnable )
      Contact( #"Dont Overwrite SP" )
   END_RUNG wire#w2
   RUNG wire#powerrail
      Contact( #inputManunalFlag )
   END_RUNG wire#w3
   RUNG wire#powerrail
      I_Contact( #notInhibited )
      Move(in := 4, out1 => #hmi.Config.mode)
      Move(in := #hmi.Config.inhibitedOutput, out1 => #hmi.Controls.manualOutput)
   END_RUNG wire#w2
   RUNG wire#powerrail
      Contact( #hmi.Status.faulted )
      Contact( #hmi.Config.allowPvFaultOverride )
      P_Trig( #triggers[1] )
   END_RUNG wire#w2
   RUNG wire#powerrail
      Contact( #hmi.Status.faulted )
      I_Contact( #hmi.Config.allowPvFaultOverride )
   END_RUNG wire#w2
   RUNG wire#w2
      S_Coil( #hmi.Controls.manualEnable )
   END_RUNG
   // the same network as SCL:
   #_w1 := #hmi.Controls.manualEnable AND NOT #trig;   // rising edge of #hmi.Controls.manualEnable
   #trig := #hmi.Controls.manualEnable;
   #_w2 := #hmi.Controls.manualEnable AND NOT #trig2;   // rising edge of #hmi.Controls.manualEnable
   #trig2 := #hmi.Controls.manualEnable;
   IF NOT #notInhibited THEN
       #hmi.Config.mode := 4;
       #hmi.Controls.manualOutput := #hmi.Config.inhibitedOutput;
   END_IF;
   #_w3 := #hmi.Status.faulted AND #hmi.Config.allowPvFaultOverride;
   #_w4 := #_w3 AND NOT #triggers[1];   // rising edge
   #triggers[1] := #_w3;
   IF ((#_w1 OR #inputManunalFlag) AND NOT #inputRemoteFlag AND NOT #hmi.Controls.remoteEnable AND NOT #"Dont Overwrite SP") OR ((#_w2 OR #inputManunalFlag) AND NOT #inputRemoteFlag AND NOT #hmi.Controls.remoteEnable AND #"Dont Overwrite SP") OR NOT #notInhibited OR #_w4 OR (#hmi.Status.faulted AND NOT #hmi.Config.allowPvFaultOverride) THEN
       #pid.ManualEnable := TRUE;
       #hmi.Controls.manualEnable := TRUE;
   END_IF;
END_REGION

